(* Logix 5000 project; controller PLC_MCC1300_75F1 vendor 1 type 14 code 166 rev 32.11; software revision 32.04; part 46 of 83 *)
(* tags used below, declared in another part *)
   GP_PosWindow : GP_PosWindow;
   M30xTrimWheel : MAC_TrimmingWheels[5];
   M30xTrimWheel_ALM : MAC_TrimmingWheels_ALM[5];
   M30xTrimWheel_HMR : MAC_TrimmingWheels_HMR[5];
   M30xTrimWheel_HMW : MAC_TrimmingWheels_HMW[5];
   TMP_dIndex : DINT;
   xAlwaysOFF : BOOL;
   xAlwaysON : BOOL;
   Z301 : MAC_Zone_ML;
(* MainProgram, continued *)

ROUTINE M30xTrimWheel_Faults   (* ladder *)
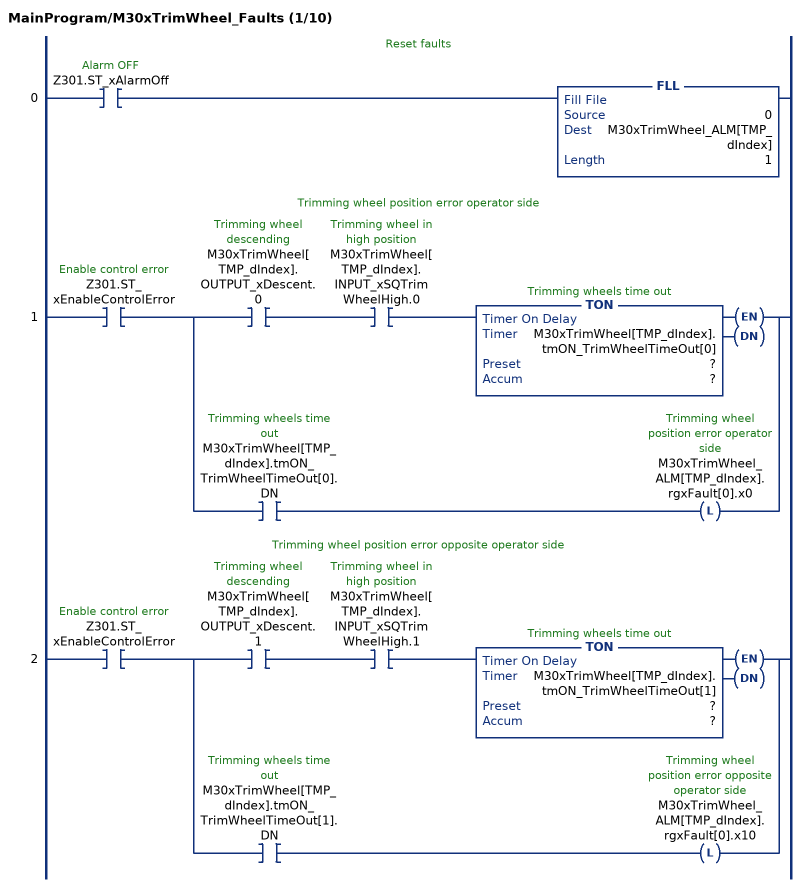
   // Reset faults
   0: XIC(Z301.ST_xAlarmOff)FLL(0,M30xTrimWheel_ALM[TMP_dIndex],1);
   // Trimming wheel position error operator side
   1: XIC(Z301.ST_xEnableControlError)[XIC(M30xTrimWheel[TMP_dIndex].OUTPUT_xDescent.0) XIC(M30xTrimWheel[TMP_dIndex].INPUT_xSQTrimWheelHigh.0) TON(M30xTrimWheel[TMP_dIndex].tmON_TrimWheelTimeOut[0],?,?) ,XIC(M30xTrimWheel[TMP_dIndex].tmON_TrimWheelTimeOut[0].DN) OTL(M30xTrimWheel_ALM[TMP_dIndex].rgxFault[0].x0) ];
   // Trimming wheel position error opposite operator side
   2: XIC(Z301.ST_xEnableControlError)[XIC(M30xTrimWheel[TMP_dIndex].OUTPUT_xDescent.1) XIC(M30xTrimWheel[TMP_dIndex].INPUT_xSQTrimWheelHigh.1) TON(M30xTrimWheel[TMP_dIndex].tmON_TrimWheelTimeOut[1],?,?) ,XIC(M30xTrimWheel[TMP_dIndex].tmON_TrimWheelTimeOut[1].DN) OTL(M30xTrimWheel_ALM[TMP_dIndex].rgxFault[0].x10) ];
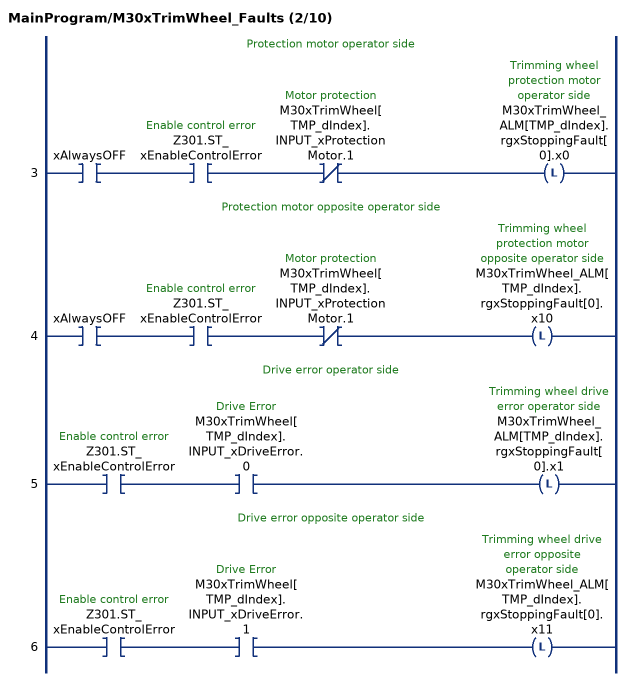
   // Protection motor operator side
   3: XIC(xAlwaysOFF)XIC(Z301.ST_xEnableControlError)XIO(M30xTrimWheel[TMP_dIndex].INPUT_xProtectionMotor.1)OTL(M30xTrimWheel_ALM[TMP_dIndex].rgxStoppingFault[0].x0);
   // Protection motor opposite operator side
   4: XIC(xAlwaysOFF)XIC(Z301.ST_xEnableControlError)XIO(M30xTrimWheel[TMP_dIndex].INPUT_xProtectionMotor.1)OTL(M30xTrimWheel_ALM[TMP_dIndex].rgxStoppingFault[0].x10);
   // Drive error operator side
   5: XIC(Z301.ST_xEnableControlError)XIC(M30xTrimWheel[TMP_dIndex].INPUT_xDriveError.0)OTL(M30xTrimWheel_ALM[TMP_dIndex].rgxStoppingFault[0].x1);
   // Drive error opposite operator side
   6: XIC(Z301.ST_xEnableControlError)XIC(M30xTrimWheel[TMP_dIndex].INPUT_xDriveError.1)OTL(M30xTrimWheel_ALM[TMP_dIndex].rgxStoppingFault[0].x11);
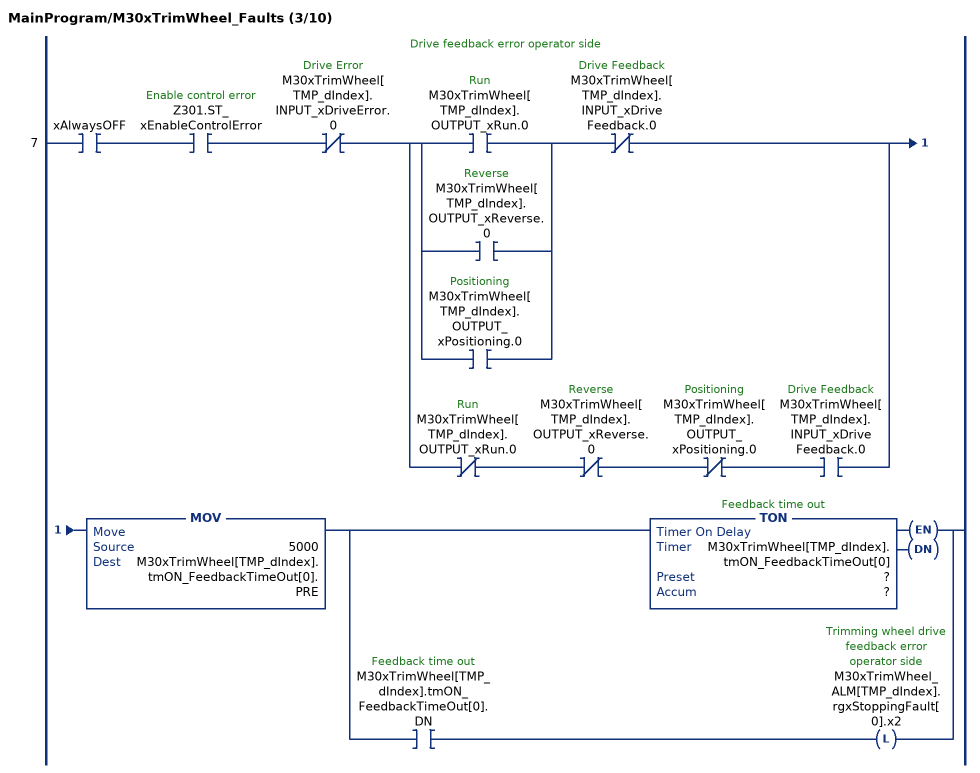
   // Drive feedback error operator side
   7: XIC(xAlwaysOFF)XIC(Z301.ST_xEnableControlError)XIO(M30xTrimWheel[TMP_dIndex].INPUT_xDriveError.0)[[XIC(M30xTrimWheel[TMP_dIndex].OUTPUT_xRun.0) ,XIC(M30xTrimWheel[TMP_dIndex].OUTPUT_xReverse.0) ,XIC(M30xTrimWheel[TMP_dIndex].OUTPUT_xPositioning.0) ] XIO(M30xTrimWheel[TMP_dIndex].INPUT_xDriveFeedback.0) ,XIO(M30xTrimWheel[TMP_dIndex].OUTPUT_xRun.0) XIO(M30xTrimWheel[TMP_dIndex].OUTPUT_xReverse.0) XIO(M30xTrimWheel[TMP_dIndex].OUTPUT_xPositioning.0) XIC(M30xTrimWheel[TMP_dIndex].INPUT_xDriveFeedback.0) ]MOV(5000,M30xTrimWheel[TMP_dIndex].tmON_FeedbackTimeOut[0].PRE)[TON(M30xTrimWheel[TMP_dIndex].tmON_FeedbackTimeOut[0],?,?) ,XIC(M30xTrimWheel[TMP_dIndex].tmON_FeedbackTimeOut[0].DN) OTL(M30xTrimWheel_ALM[TMP_dIndex].rgxStoppingFault[0].x2) ];
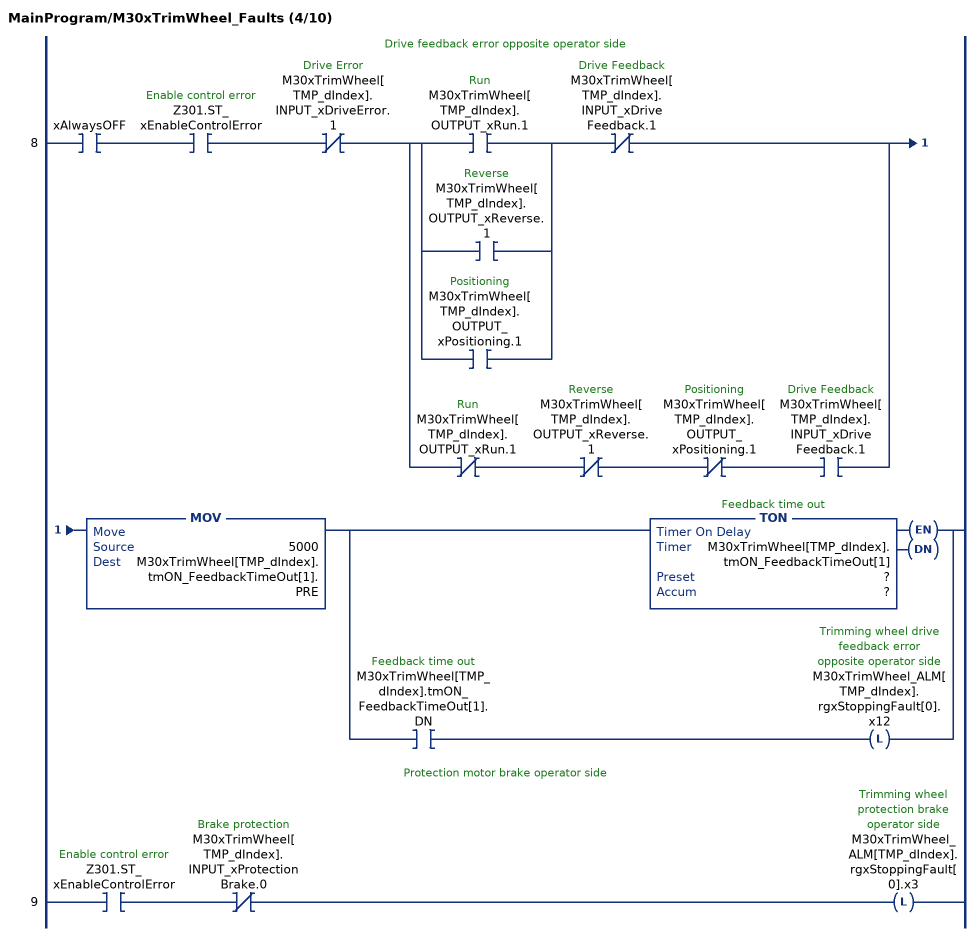
   // Drive feedback error opposite operator side
   8: XIC(xAlwaysOFF)XIC(Z301.ST_xEnableControlError)XIO(M30xTrimWheel[TMP_dIndex].INPUT_xDriveError.1)[[XIC(M30xTrimWheel[TMP_dIndex].OUTPUT_xRun.1) ,XIC(M30xTrimWheel[TMP_dIndex].OUTPUT_xReverse.1) ,XIC(M30xTrimWheel[TMP_dIndex].OUTPUT_xPositioning.1) ] XIO(M30xTrimWheel[TMP_dIndex].INPUT_xDriveFeedback.1) ,XIO(M30xTrimWheel[TMP_dIndex].OUTPUT_xRun.1) XIO(M30xTrimWheel[TMP_dIndex].OUTPUT_xReverse.1) XIO(M30xTrimWheel[TMP_dIndex].OUTPUT_xPositioning.1) XIC(M30xTrimWheel[TMP_dIndex].INPUT_xDriveFeedback.1) ]MOV(5000,M30xTrimWheel[TMP_dIndex].tmON_FeedbackTimeOut[1].PRE)[TON(M30xTrimWheel[TMP_dIndex].tmON_FeedbackTimeOut[1],?,?) ,XIC(M30xTrimWheel[TMP_dIndex].tmON_FeedbackTimeOut[1].DN) OTL(M30xTrimWheel_ALM[TMP_dIndex].rgxStoppingFault[0].x12) ];
   // Protection motor brake operator side
   9: XIC(Z301.ST_xEnableControlError)XIO(M30xTrimWheel[TMP_dIndex].INPUT_xProtectionBrake.0)OTL(M30xTrimWheel_ALM[TMP_dIndex].rgxStoppingFault[0].x3);
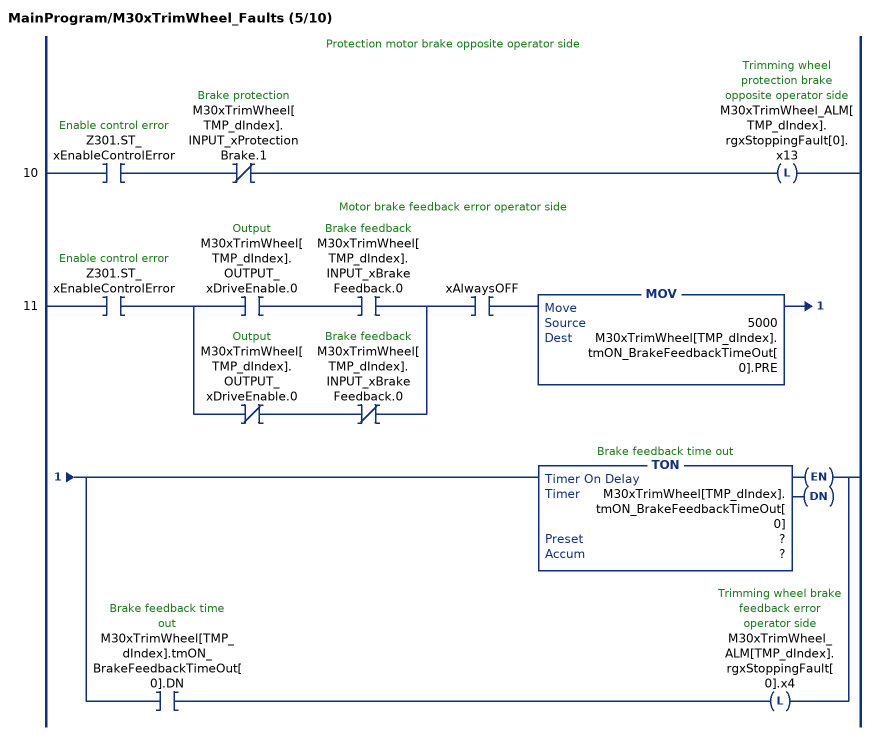
   // Protection motor brake opposite operator side
   10: XIC(Z301.ST_xEnableControlError)XIO(M30xTrimWheel[TMP_dIndex].INPUT_xProtectionBrake.1)OTL(M30xTrimWheel_ALM[TMP_dIndex].rgxStoppingFault[0].x13);
   // Motor brake feedback error operator side
   11: XIC(Z301.ST_xEnableControlError)[XIC(M30xTrimWheel[TMP_dIndex].OUTPUT_xDriveEnable.0) XIC(M30xTrimWheel[TMP_dIndex].INPUT_xBrakeFeedback.0) ,XIO(M30xTrimWheel[TMP_dIndex].OUTPUT_xDriveEnable.0) XIO(M30xTrimWheel[TMP_dIndex].INPUT_xBrakeFeedback.0) ]XIC(xAlwaysOFF)MOV(5000,M30xTrimWheel[TMP_dIndex].tmON_BrakeFeedbackTimeOut[0].PRE)[TON(M30xTrimWheel[TMP_dIndex].tmON_BrakeFeedbackTimeOut[0],?,?) ,XIC(M30xTrimWheel[TMP_dIndex].tmON_BrakeFeedbackTimeOut[0].DN) OTL(M30xTrimWheel_ALM[TMP_dIndex].rgxStoppingFault[0].x4) ];
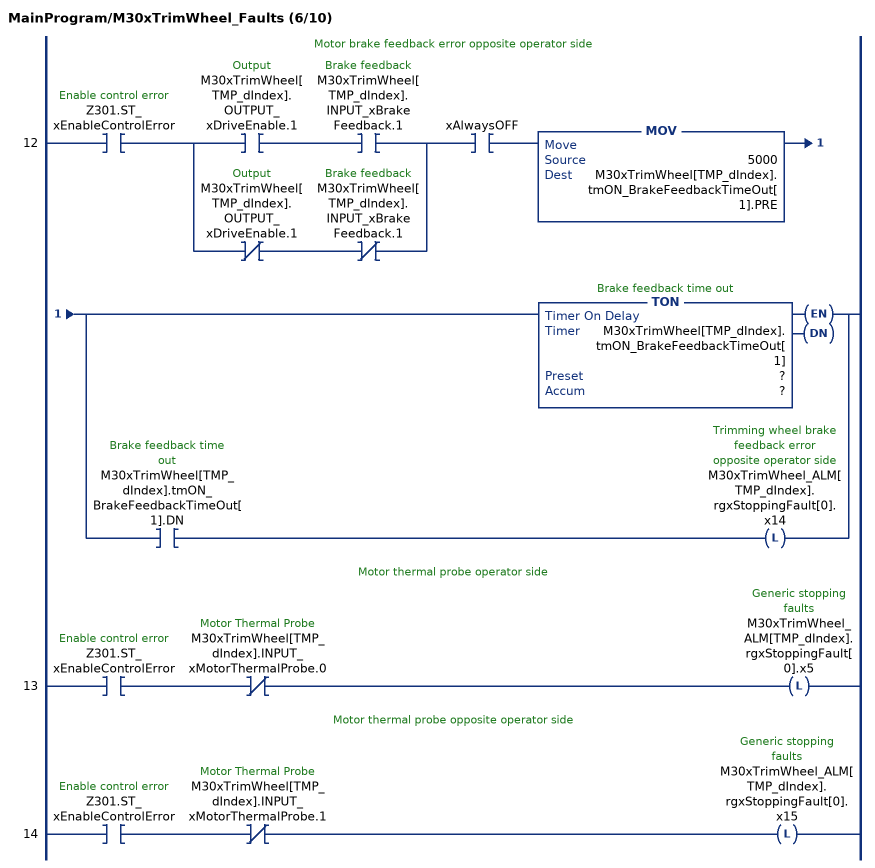
   // Motor brake feedback error opposite operator side
   12: XIC(Z301.ST_xEnableControlError)[XIC(M30xTrimWheel[TMP_dIndex].OUTPUT_xDriveEnable.1) XIC(M30xTrimWheel[TMP_dIndex].INPUT_xBrakeFeedback.1) ,XIO(M30xTrimWheel[TMP_dIndex].OUTPUT_xDriveEnable.1) XIO(M30xTrimWheel[TMP_dIndex].INPUT_xBrakeFeedback.1) ]XIC(xAlwaysOFF)MOV(5000,M30xTrimWheel[TMP_dIndex].tmON_BrakeFeedbackTimeOut[1].PRE)[TON(M30xTrimWheel[TMP_dIndex].tmON_BrakeFeedbackTimeOut[1],?,?) ,XIC(M30xTrimWheel[TMP_dIndex].tmON_BrakeFeedbackTimeOut[1].DN) OTL(M30xTrimWheel_ALM[TMP_dIndex].rgxStoppingFault[0].x14) ];
   // Motor thermal probe operator side
   13: XIC(Z301.ST_xEnableControlError)XIO(M30xTrimWheel[TMP_dIndex].INPUT_xMotorThermalProbe.0)OTL(M30xTrimWheel_ALM[TMP_dIndex].rgxStoppingFault[0].x5);
   // Motor thermal probe opposite operator side
   14: XIC(Z301.ST_xEnableControlError)XIO(M30xTrimWheel[TMP_dIndex].INPUT_xMotorThermalProbe.1)OTL(M30xTrimWheel_ALM[TMP_dIndex].rgxStoppingFault[0].x15);
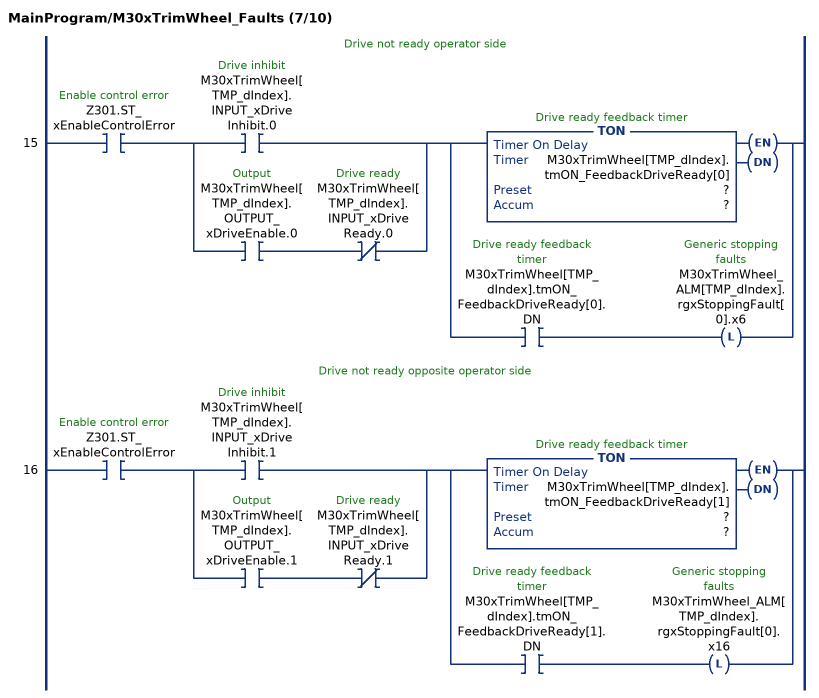
   // Drive not ready operator side
   15: XIC(Z301.ST_xEnableControlError)[XIC(M30xTrimWheel[TMP_dIndex].INPUT_xDriveInhibit.0) ,XIC(M30xTrimWheel[TMP_dIndex].OUTPUT_xDriveEnable.0) XIO(M30xTrimWheel[TMP_dIndex].INPUT_xDriveReady.0) ][TON(M30xTrimWheel[TMP_dIndex].tmON_FeedbackDriveReady[0],?,?) ,XIC(M30xTrimWheel[TMP_dIndex].tmON_FeedbackDriveReady[0].DN) OTL(M30xTrimWheel_ALM[TMP_dIndex].rgxStoppingFault[0].x6) ];
   // Drive not ready opposite operator side
   16: XIC(Z301.ST_xEnableControlError)[XIC(M30xTrimWheel[TMP_dIndex].INPUT_xDriveInhibit.1) ,XIC(M30xTrimWheel[TMP_dIndex].OUTPUT_xDriveEnable.1) XIO(M30xTrimWheel[TMP_dIndex].INPUT_xDriveReady.1) ][TON(M30xTrimWheel[TMP_dIndex].tmON_FeedbackDriveReady[1],?,?) ,XIC(M30xTrimWheel[TMP_dIndex].tmON_FeedbackDriveReady[1].DN) OTL(M30xTrimWheel_ALM[TMP_dIndex].rgxStoppingFault[0].x16) ];
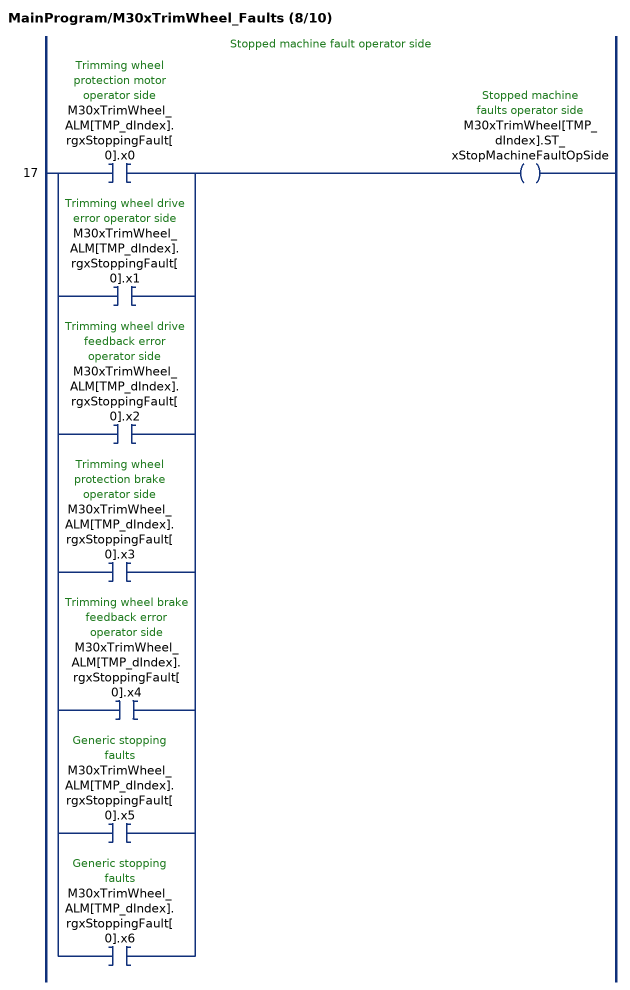
   // Stopped machine fault operator side
   17: [XIC(M30xTrimWheel_ALM[TMP_dIndex].rgxStoppingFault[0].x0) ,XIC(M30xTrimWheel_ALM[TMP_dIndex].rgxStoppingFault[0].x1) ,XIC(M30xTrimWheel_ALM[TMP_dIndex].rgxStoppingFault[0].x2) ,XIC(M30xTrimWheel_ALM[TMP_dIndex].rgxStoppingFault[0].x3) ,XIC(M30xTrimWheel_ALM[TMP_dIndex].rgxStoppingFault[0].x4) ,XIC(M30xTrimWheel_ALM[TMP_dIndex].rgxStoppingFault[0].x5) ,XIC(M30xTrimWheel_ALM[TMP_dIndex].rgxStoppingFault[0].x6) ]OTE(M30xTrimWheel[TMP_dIndex].ST_xStopMachineFaultOpSide);
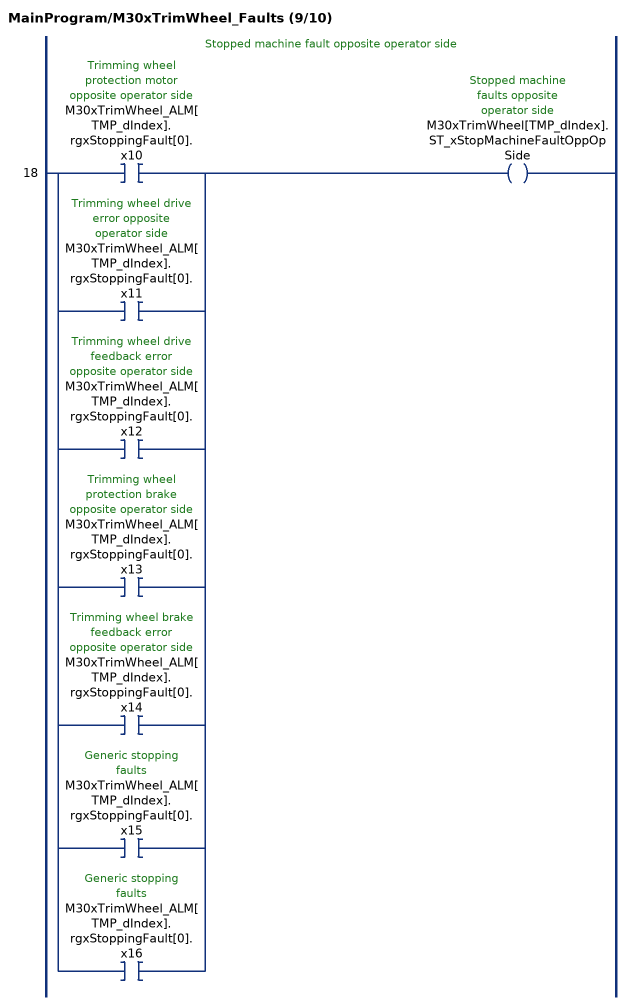
   // Stopped machine fault opposite operator side
   18: [XIC(M30xTrimWheel_ALM[TMP_dIndex].rgxStoppingFault[0].x10) ,XIC(M30xTrimWheel_ALM[TMP_dIndex].rgxStoppingFault[0].x11) ,XIC(M30xTrimWheel_ALM[TMP_dIndex].rgxStoppingFault[0].x12) ,XIC(M30xTrimWheel_ALM[TMP_dIndex].rgxStoppingFault[0].x13) ,XIC(M30xTrimWheel_ALM[TMP_dIndex].rgxStoppingFault[0].x14) ,XIC(M30xTrimWheel_ALM[TMP_dIndex].rgxStoppingFault[0].x15) ,XIC(M30xTrimWheel_ALM[TMP_dIndex].rgxStoppingFault[0].x16) ]OTE(M30xTrimWheel[TMP_dIndex].ST_xStopMachineFaultOppOpSide);
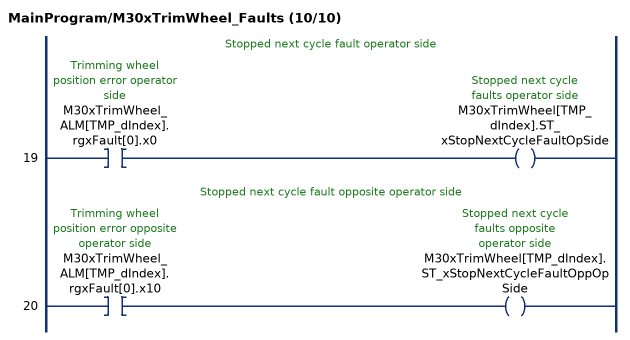
   // Stopped next cycle fault operator side
   19: XIC(M30xTrimWheel_ALM[TMP_dIndex].rgxFault[0].x0)OTE(M30xTrimWheel[TMP_dIndex].ST_xStopNextCycleFaultOpSide);
   // Stopped next cycle fault opposite operator side
   20: XIC(M30xTrimWheel_ALM[TMP_dIndex].rgxFault[0].x10)OTE(M30xTrimWheel[TMP_dIndex].ST_xStopNextCycleFaultOppOpSide);
END_ROUTINE

ROUTINE M30xTrimWheel_Logic   (* ladder *)
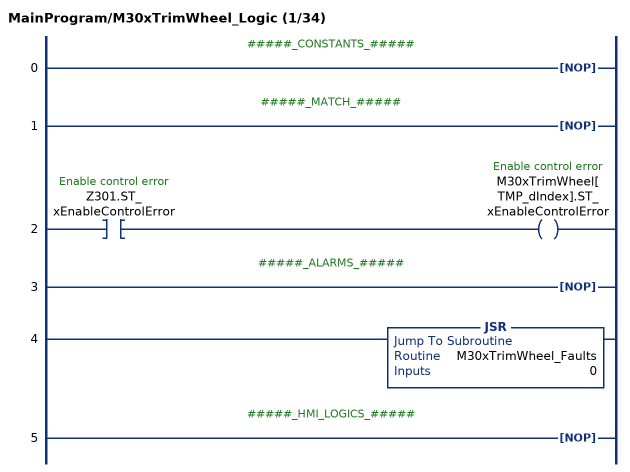
   // #####_CONSTANTS_#####
   0: NOP();
   // #####_MATCH_#####
   1: NOP();
   2: XIC(Z301.ST_xEnableControlError)OTE(M30xTrimWheel[TMP_dIndex].ST_xEnableControlError);
   // #####_ALARMS_#####
   3: NOP();
   4: JSR(M30xTrimWheel_Faults,0);
   // #####_HMI_LOGICS_#####
   5: NOP();
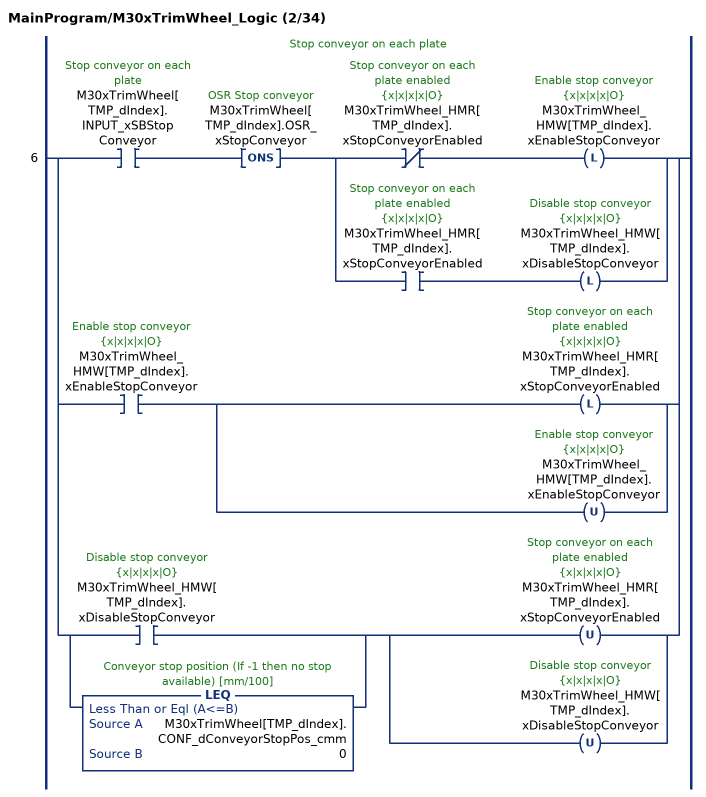
   // Stop conveyor on each plate
   6: [XIC(M30xTrimWheel[TMP_dIndex].INPUT_xSBStopConveyor) ONS(M30xTrimWheel[TMP_dIndex].OSR_xStopConveyor) [XIO(M30xTrimWheel_HMR[TMP_dIndex].xStopConveyorEnabled) OTL(M30xTrimWheel_HMW[TMP_dIndex].xEnableStopConveyor) ,XIC(M30xTrimWheel_HMR[TMP_dIndex].xStopConveyorEnabled) OTL(M30xTrimWheel_HMW[TMP_dIndex].xDisableStopConveyor) ] ,[XIC(M30xTrimWheel_HMW[TMP_dIndex].xEnableStopConveyor) [OTL(M30xTrimWheel_HMR[TMP_dIndex].xStopConveyorEnabled) ,OTU(M30xTrimWheel_HMW[TMP_dIndex].xEnableStopConveyor) ] ,[XIC(M30xTrimWheel_HMW[TMP_dIndex].xDisableStopConveyor) ,LEQ(M30xTrimWheel[TMP_dIndex].CONF_dConveyorStopPos_cmm,0) ] [OTU(M30xTrimWheel_HMR[TMP_dIndex].xStopConveyorEnabled) ,OTU(M30xTrimWheel_HMW[TMP_dIndex].xDisableStopConveyor) ] ] ];
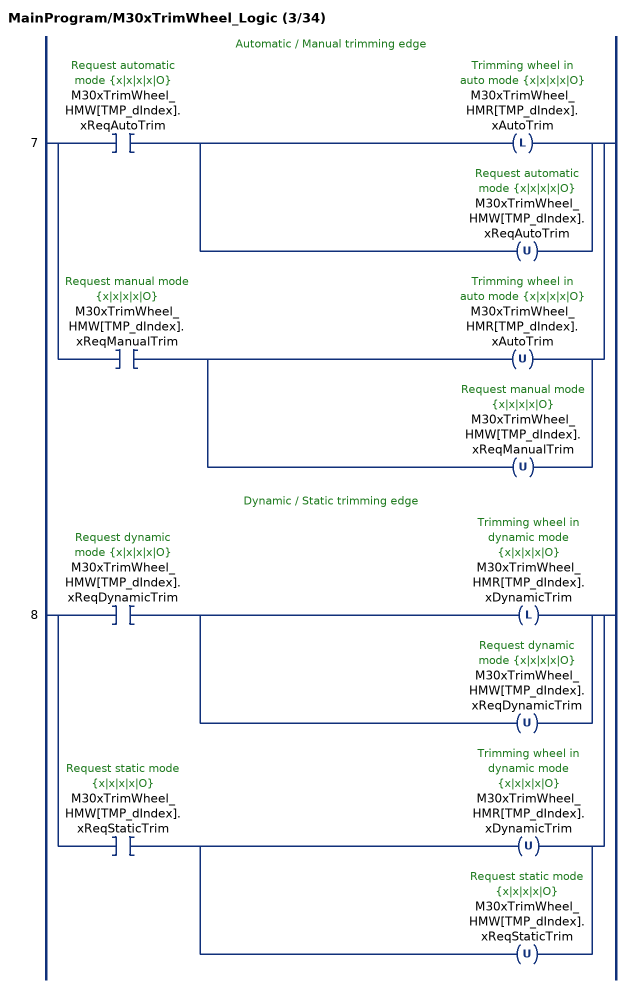
   // Automatic / Manual trimming edge
   7: [XIC(M30xTrimWheel_HMW[TMP_dIndex].xReqAutoTrim) [OTL(M30xTrimWheel_HMR[TMP_dIndex].xAutoTrim) ,OTU(M30xTrimWheel_HMW[TMP_dIndex].xReqAutoTrim) ] ,XIC(M30xTrimWheel_HMW[TMP_dIndex].xReqManualTrim) [OTU(M30xTrimWheel_HMR[TMP_dIndex].xAutoTrim) ,OTU(M30xTrimWheel_HMW[TMP_dIndex].xReqManualTrim) ] ];
   // Dynamic / Static trimming edge
   8: [XIC(M30xTrimWheel_HMW[TMP_dIndex].xReqDynamicTrim) [OTL(M30xTrimWheel_HMR[TMP_dIndex].xDynamicTrim) ,OTU(M30xTrimWheel_HMW[TMP_dIndex].xReqDynamicTrim) ] ,XIC(M30xTrimWheel_HMW[TMP_dIndex].xReqStaticTrim) [OTU(M30xTrimWheel_HMR[TMP_dIndex].xDynamicTrim) ,OTU(M30xTrimWheel_HMW[TMP_dIndex].xReqStaticTrim) ] ];
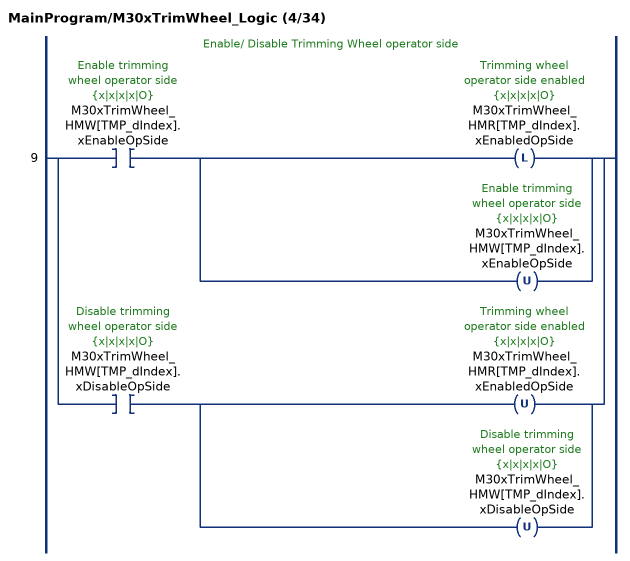
   // Enable/ Disable Trimming Wheel operator side
   9: [XIC(M30xTrimWheel_HMW[TMP_dIndex].xEnableOpSide) [OTL(M30xTrimWheel_HMR[TMP_dIndex].xEnabledOpSide) ,OTU(M30xTrimWheel_HMW[TMP_dIndex].xEnableOpSide) ] ,XIC(M30xTrimWheel_HMW[TMP_dIndex].xDisableOpSide) [OTU(M30xTrimWheel_HMR[TMP_dIndex].xEnabledOpSide) ,OTU(M30xTrimWheel_HMW[TMP_dIndex].xDisableOpSide) ] ];
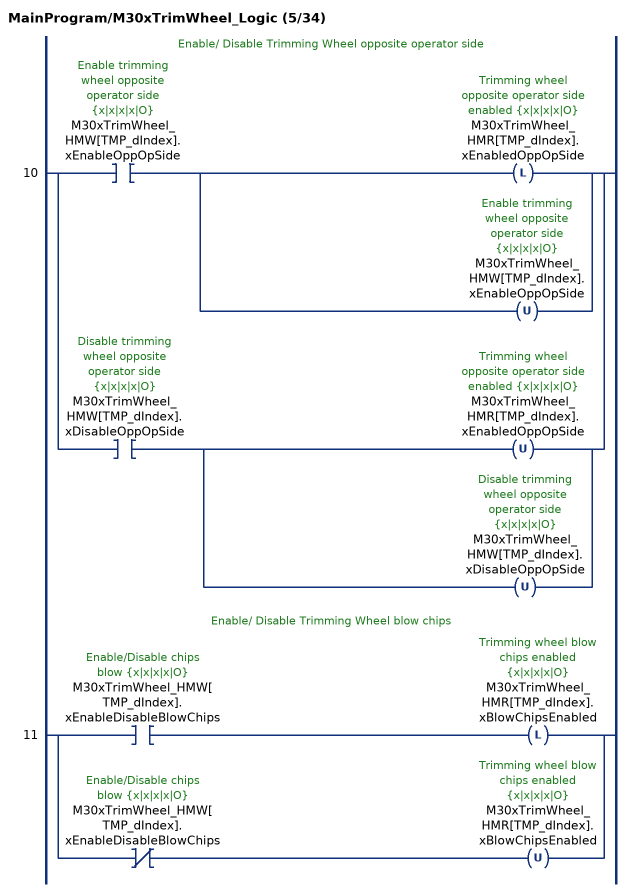
   // Enable/ Disable Trimming Wheel opposite operator side
   10: [XIC(M30xTrimWheel_HMW[TMP_dIndex].xEnableOppOpSide) [OTL(M30xTrimWheel_HMR[TMP_dIndex].xEnabledOppOpSide) ,OTU(M30xTrimWheel_HMW[TMP_dIndex].xEnableOppOpSide) ] ,XIC(M30xTrimWheel_HMW[TMP_dIndex].xDisableOppOpSide) [OTU(M30xTrimWheel_HMR[TMP_dIndex].xEnabledOppOpSide) ,OTU(M30xTrimWheel_HMW[TMP_dIndex].xDisableOppOpSide) ] ];
   // Enable/ Disable Trimming Wheel blow chips
   11: [XIC(M30xTrimWheel_HMW[TMP_dIndex].xEnableDisableBlowChips) OTL(M30xTrimWheel_HMR[TMP_dIndex].xBlowChipsEnabled) ,XIO(M30xTrimWheel_HMW[TMP_dIndex].xEnableDisableBlowChips) OTU(M30xTrimWheel_HMR[TMP_dIndex].xBlowChipsEnabled) ];
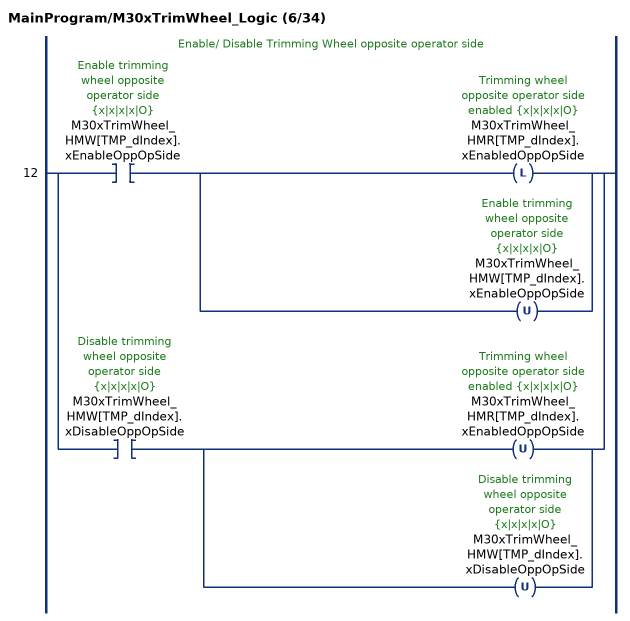
   // Enable/ Disable Trimming Wheel opposite operator side
   12: [XIC(M30xTrimWheel_HMW[TMP_dIndex].xEnableOppOpSide) [OTL(M30xTrimWheel_HMR[TMP_dIndex].xEnabledOppOpSide) ,OTU(M30xTrimWheel_HMW[TMP_dIndex].xEnableOppOpSide) ] ,XIC(M30xTrimWheel_HMW[TMP_dIndex].xDisableOppOpSide) [OTU(M30xTrimWheel_HMR[TMP_dIndex].xEnabledOppOpSide) ,OTU(M30xTrimWheel_HMW[TMP_dIndex].xDisableOppOpSide) ] ];
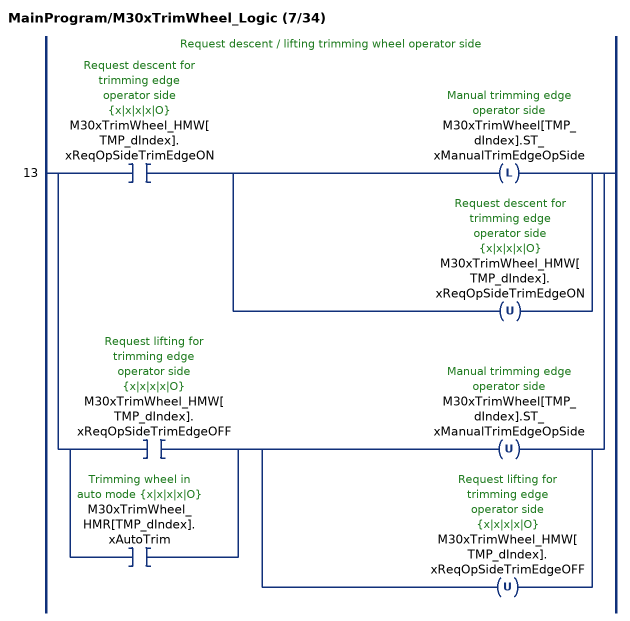
   // Request descent / lifting trimming wheel operator side
   13: [XIC(M30xTrimWheel_HMW[TMP_dIndex].xReqOpSideTrimEdgeON) [OTL(M30xTrimWheel[TMP_dIndex].ST_xManualTrimEdgeOpSide) ,OTU(M30xTrimWheel_HMW[TMP_dIndex].xReqOpSideTrimEdgeON) ] ,[XIC(M30xTrimWheel_HMW[TMP_dIndex].xReqOpSideTrimEdgeOFF) ,XIC(M30xTrimWheel_HMR[TMP_dIndex].xAutoTrim) ] [OTU(M30xTrimWheel[TMP_dIndex].ST_xManualTrimEdgeOpSide) ,OTU(M30xTrimWheel_HMW[TMP_dIndex].xReqOpSideTrimEdgeOFF) ] ];
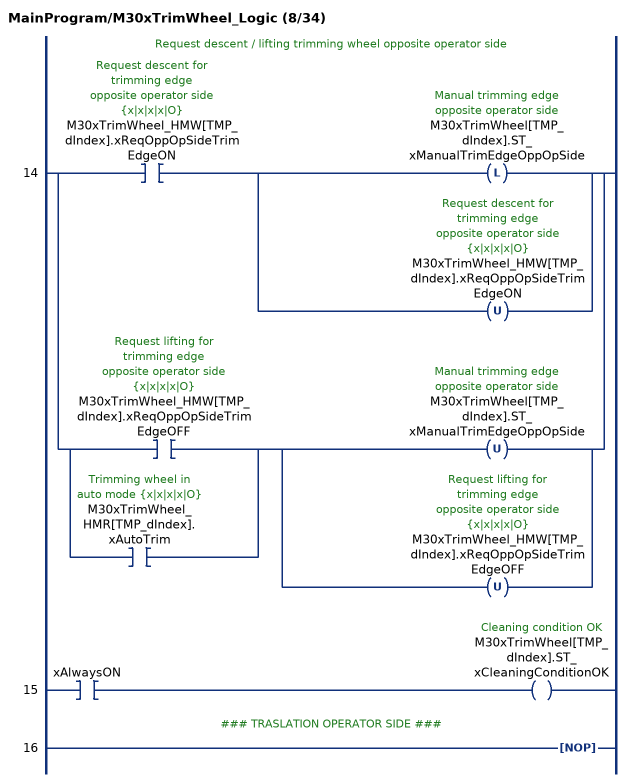
   // Request descent / lifting trimming wheel opposite operator side
   14: [XIC(M30xTrimWheel_HMW[TMP_dIndex].xReqOppOpSideTrimEdgeON) [OTL(M30xTrimWheel[TMP_dIndex].ST_xManualTrimEdgeOppOpSide) ,OTU(M30xTrimWheel_HMW[TMP_dIndex].xReqOppOpSideTrimEdgeON) ] ,[XIC(M30xTrimWheel_HMW[TMP_dIndex].xReqOppOpSideTrimEdgeOFF) ,XIC(M30xTrimWheel_HMR[TMP_dIndex].xAutoTrim) ] [OTU(M30xTrimWheel[TMP_dIndex].ST_xManualTrimEdgeOppOpSide) ,OTU(M30xTrimWheel_HMW[TMP_dIndex].xReqOppOpSideTrimEdgeOFF) ] ];
   15: XIC(xAlwaysON)OTE(M30xTrimWheel[TMP_dIndex].ST_xCleaningConditionOK);
   // ### TRASLATION OPERATOR SIDE ###
   16: NOP();
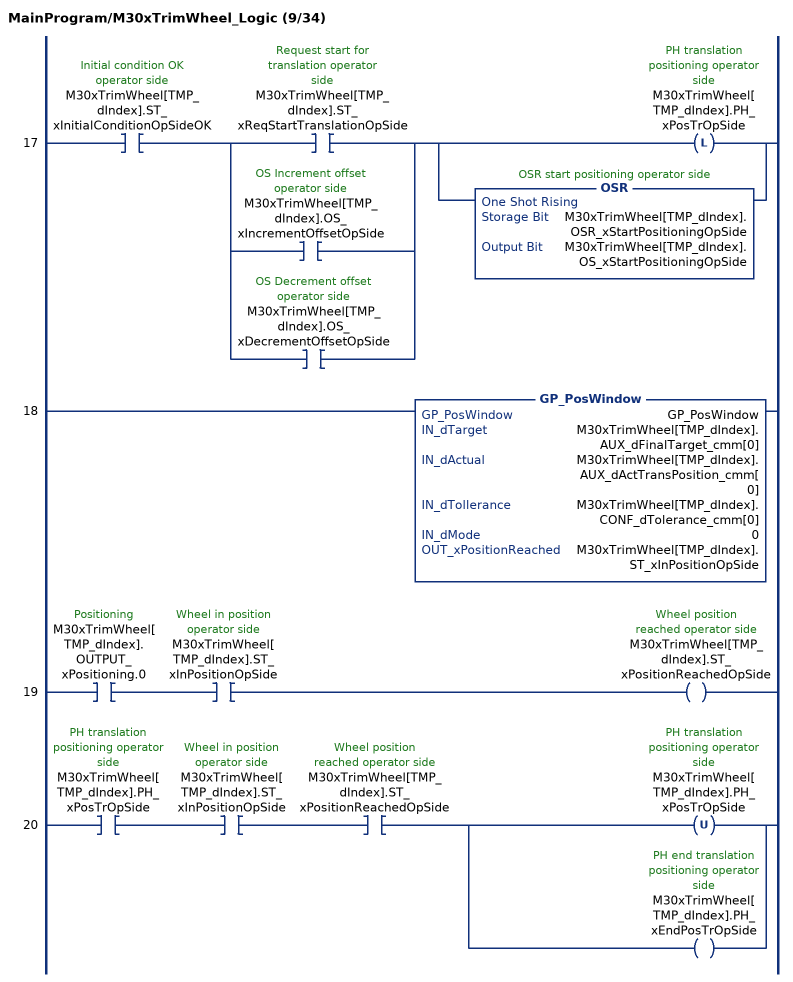
   17: XIC(M30xTrimWheel[TMP_dIndex].ST_xInitialConditionOpSideOK)[XIC(M30xTrimWheel[TMP_dIndex].ST_xReqStartTranslationOpSide) ,[XIC(M30xTrimWheel[TMP_dIndex].OS_xIncrementOffsetOpSide) ,XIC(M30xTrimWheel[TMP_dIndex].OS_xDecrementOffsetOpSide) ] ][OTL(M30xTrimWheel[TMP_dIndex].PH_xPosTrOpSide) ,OSR(M30xTrimWheel[TMP_dIndex].OSR_xStartPositioningOpSide,M30xTrimWheel[TMP_dIndex].OS_xStartPositioningOpSide) ];
   18: GP_PosWindow(GP_PosWindow,M30xTrimWheel[TMP_dIndex].AUX_dFinalTarget_cmm[0],M30xTrimWheel[TMP_dIndex].AUX_dActTransPosition_cmm[0],M30xTrimWheel[TMP_dIndex].CONF_dTolerance_cmm[0],0,M30xTrimWheel[TMP_dIndex].ST_xInPositionOpSide);
   19: XIC(M30xTrimWheel[TMP_dIndex].OUTPUT_xPositioning.0)XIC(M30xTrimWheel[TMP_dIndex].ST_xInPositionOpSide)OTE(M30xTrimWheel[TMP_dIndex].ST_xPositionReachedOpSide);
   20: XIC(M30xTrimWheel[TMP_dIndex].PH_xPosTrOpSide)XIC(M30xTrimWheel[TMP_dIndex].ST_xInPositionOpSide)XIC(M30xTrimWheel[TMP_dIndex].ST_xPositionReachedOpSide)[OTU(M30xTrimWheel[TMP_dIndex].PH_xPosTrOpSide) ,OTE(M30xTrimWheel[TMP_dIndex].PH_xEndPosTrOpSide) ];
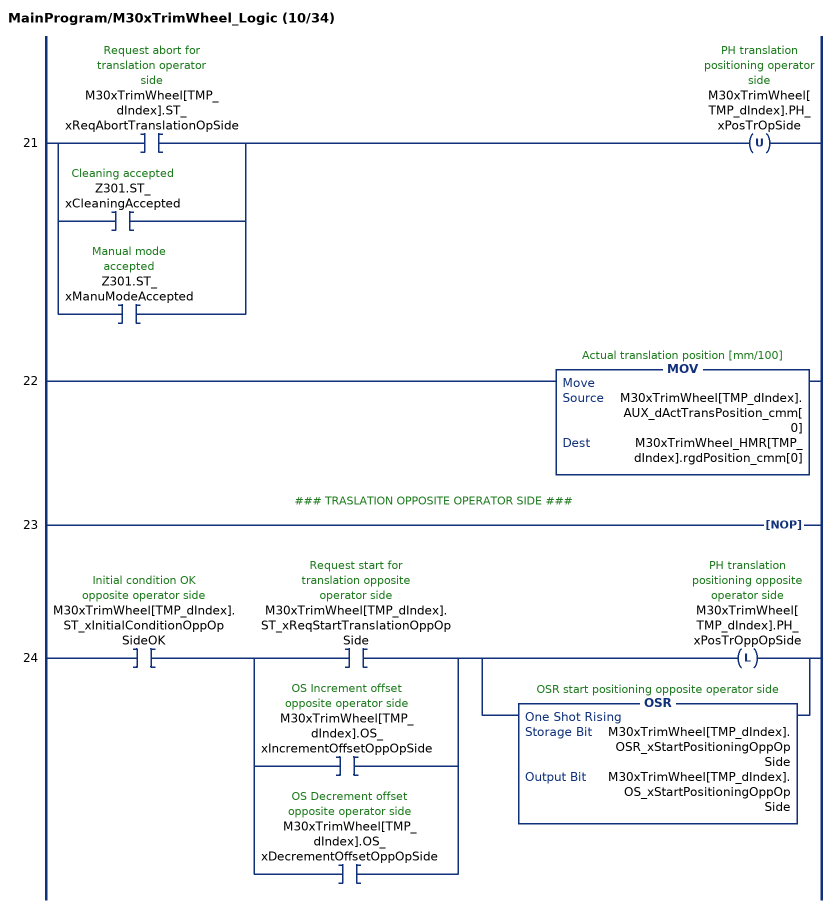
   21: [XIC(M30xTrimWheel[TMP_dIndex].ST_xReqAbortTranslationOpSide) ,XIC(Z301.ST_xCleaningAccepted) ,XIC(Z301.ST_xManuModeAccepted) ]OTU(M30xTrimWheel[TMP_dIndex].PH_xPosTrOpSide);
   22: MOV(M30xTrimWheel[TMP_dIndex].AUX_dActTransPosition_cmm[0],M30xTrimWheel_HMR[TMP_dIndex].rgdPosition_cmm[0]);
   // ### TRASLATION OPPOSITE OPERATOR SIDE ###
   23: NOP();
   24: XIC(M30xTrimWheel[TMP_dIndex].ST_xInitialConditionOppOpSideOK)[XIC(M30xTrimWheel[TMP_dIndex].ST_xReqStartTranslationOppOpSide) ,[XIC(M30xTrimWheel[TMP_dIndex].OS_xIncrementOffsetOppOpSide) ,XIC(M30xTrimWheel[TMP_dIndex].OS_xDecrementOffsetOppOpSide) ] ][OTL(M30xTrimWheel[TMP_dIndex].PH_xPosTrOppOpSide) ,OSR(M30xTrimWheel[TMP_dIndex].OSR_xStartPositioningOppOpSide,M30xTrimWheel[TMP_dIndex].OS_xStartPositioningOppOpSide) ];
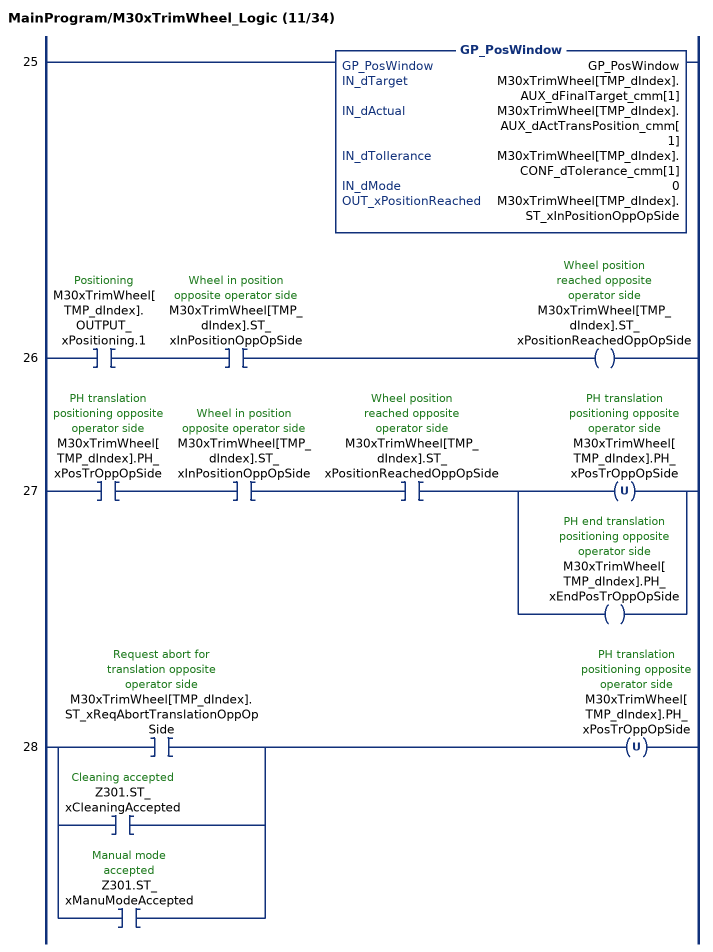
   25: GP_PosWindow(GP_PosWindow,M30xTrimWheel[TMP_dIndex].AUX_dFinalTarget_cmm[1],M30xTrimWheel[TMP_dIndex].AUX_dActTransPosition_cmm[1],M30xTrimWheel[TMP_dIndex].CONF_dTolerance_cmm[1],0,M30xTrimWheel[TMP_dIndex].ST_xInPositionOppOpSide);
   26: XIC(M30xTrimWheel[TMP_dIndex].OUTPUT_xPositioning.1)XIC(M30xTrimWheel[TMP_dIndex].ST_xInPositionOppOpSide)OTE(M30xTrimWheel[TMP_dIndex].ST_xPositionReachedOppOpSide);
   27: XIC(M30xTrimWheel[TMP_dIndex].PH_xPosTrOppOpSide)XIC(M30xTrimWheel[TMP_dIndex].ST_xInPositionOppOpSide)XIC(M30xTrimWheel[TMP_dIndex].ST_xPositionReachedOppOpSide)[OTU(M30xTrimWheel[TMP_dIndex].PH_xPosTrOppOpSide) ,OTE(M30xTrimWheel[TMP_dIndex].PH_xEndPosTrOppOpSide) ];
   28: [XIC(M30xTrimWheel[TMP_dIndex].ST_xReqAbortTranslationOppOpSide) ,XIC(Z301.ST_xCleaningAccepted) ,XIC(Z301.ST_xManuModeAccepted) ]OTU(M30xTrimWheel[TMP_dIndex].PH_xPosTrOppOpSide);
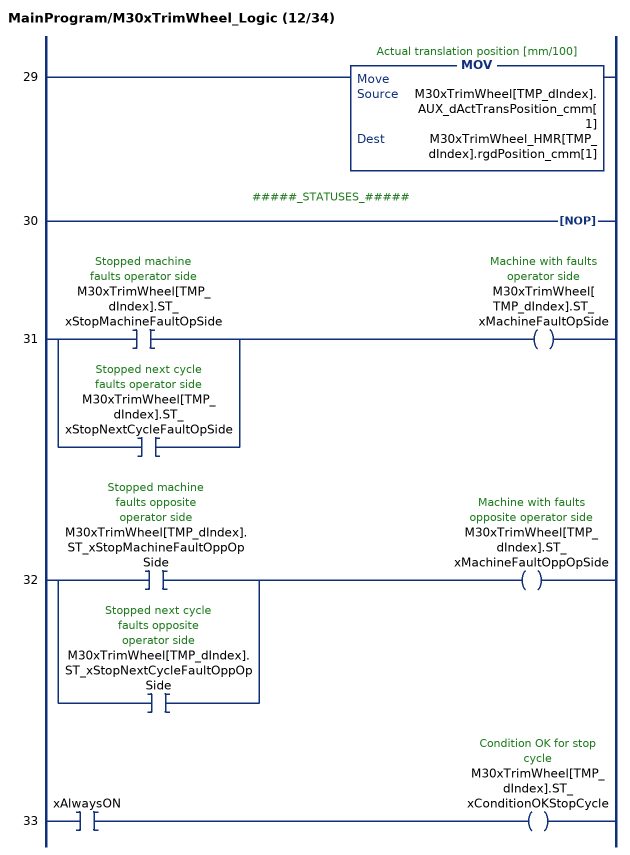
   29: MOV(M30xTrimWheel[TMP_dIndex].AUX_dActTransPosition_cmm[1],M30xTrimWheel_HMR[TMP_dIndex].rgdPosition_cmm[1]);
   // #####_STATUSES_#####
   30: NOP();
   31: [XIC(M30xTrimWheel[TMP_dIndex].ST_xStopMachineFaultOpSide) ,XIC(M30xTrimWheel[TMP_dIndex].ST_xStopNextCycleFaultOpSide) ]OTE(M30xTrimWheel[TMP_dIndex].ST_xMachineFaultOpSide);
   32: [XIC(M30xTrimWheel[TMP_dIndex].ST_xStopMachineFaultOppOpSide) ,XIC(M30xTrimWheel[TMP_dIndex].ST_xStopNextCycleFaultOppOpSide) ]OTE(M30xTrimWheel[TMP_dIndex].ST_xMachineFaultOppOpSide);
   33: XIC(xAlwaysON)OTE(M30xTrimWheel[TMP_dIndex].ST_xConditionOKStopCycle);
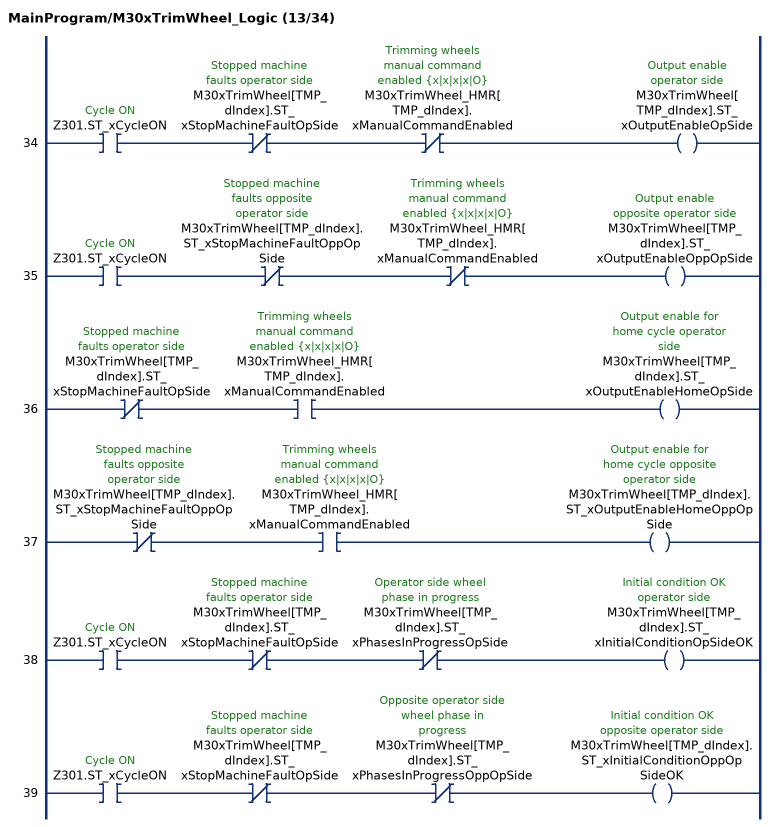
   34: XIC(Z301.ST_xCycleON)XIO(M30xTrimWheel[TMP_dIndex].ST_xStopMachineFaultOpSide)XIO(M30xTrimWheel_HMR[TMP_dIndex].xManualCommandEnabled)OTE(M30xTrimWheel[TMP_dIndex].ST_xOutputEnableOpSide);
   35: XIC(Z301.ST_xCycleON)XIO(M30xTrimWheel[TMP_dIndex].ST_xStopMachineFaultOppOpSide)XIO(M30xTrimWheel_HMR[TMP_dIndex].xManualCommandEnabled)OTE(M30xTrimWheel[TMP_dIndex].ST_xOutputEnableOppOpSide);
   36: XIO(M30xTrimWheel[TMP_dIndex].ST_xStopMachineFaultOpSide)XIC(M30xTrimWheel_HMR[TMP_dIndex].xManualCommandEnabled)OTE(M30xTrimWheel[TMP_dIndex].ST_xOutputEnableHomeOpSide);
   37: XIO(M30xTrimWheel[TMP_dIndex].ST_xStopMachineFaultOppOpSide)XIC(M30xTrimWheel_HMR[TMP_dIndex].xManualCommandEnabled)OTE(M30xTrimWheel[TMP_dIndex].ST_xOutputEnableHomeOppOpSide);
   38: XIC(Z301.ST_xCycleON)XIO(M30xTrimWheel[TMP_dIndex].ST_xStopMachineFaultOpSide)XIO(M30xTrimWheel[TMP_dIndex].ST_xPhasesInProgressOpSide)OTE(M30xTrimWheel[TMP_dIndex].ST_xInitialConditionOpSideOK);
   39: XIC(Z301.ST_xCycleON)XIO(M30xTrimWheel[TMP_dIndex].ST_xStopMachineFaultOpSide)XIO(M30xTrimWheel[TMP_dIndex].ST_xPhasesInProgressOppOpSide)OTE(M30xTrimWheel[TMP_dIndex].ST_xInitialConditionOppOpSideOK);
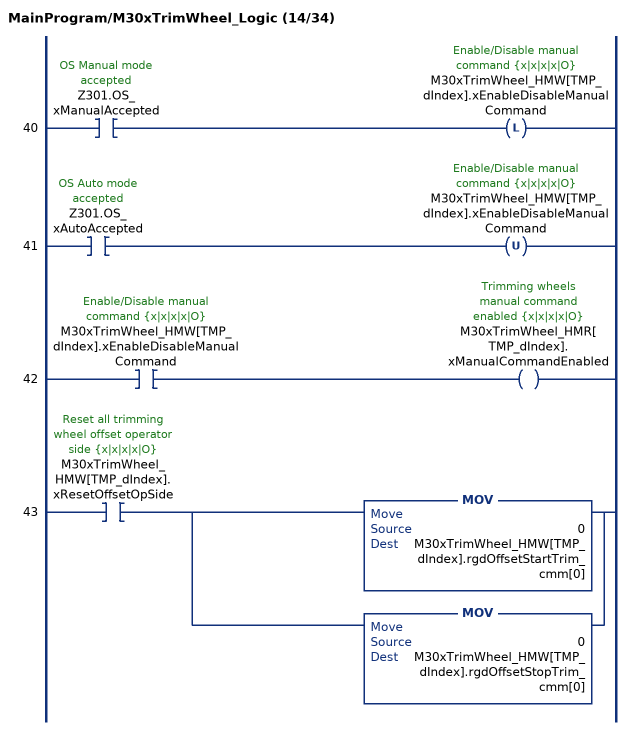
   40: XIC(Z301.OS_xManualAccepted)OTL(M30xTrimWheel_HMW[TMP_dIndex].xEnableDisableManualCommand);
   41: XIC(Z301.OS_xAutoAccepted)OTU(M30xTrimWheel_HMW[TMP_dIndex].xEnableDisableManualCommand);
   42: XIC(M30xTrimWheel_HMW[TMP_dIndex].xEnableDisableManualCommand)OTE(M30xTrimWheel_HMR[TMP_dIndex].xManualCommandEnabled);
   43: XIC(M30xTrimWheel_HMW[TMP_dIndex].xResetOffsetOpSide)[MOV(0,M30xTrimWheel_HMW[TMP_dIndex].rgdOffsetStartTrim_cmm[0]) ,MOV(0,M30xTrimWheel_HMW[TMP_dIndex].rgdOffsetStopTrim_cmm[0]) ];
